// TIA Portal project "Automatizare_RT" (V17)

(* hardware
DEVICE "S7-300/ET200M station_1"  S7-300 station
   slot 0: "Rail_0"  Rail  6ES7 390-1***0-0AA0
   slot 1: "PS 307 5A_1"  PS 307 5A  6ES7 307-1EA00-0AA0
   slot 2: "PLC_1"  CPU 319-3 PN/DP  6ES7 318-3EL00-0AB0  V2.6
      slot 1: "MPI/DP interface_1"  X1
      slot 2: "DP interface_1"  X2
      slot 3: "PROFINET interface_1"  PN-IO
         slot 1: "Port_1"  Port
   slot 4: "DI 8/DO 8x24VDC/0.5A_1"  DI8/DO8 x 24VDC / 0.5A  6ES7 323-1BH01-0AA0
   slot 5: "DI 8/DO 8x24VDC/0.5A_2"  DI8/DO8 x 24VDC / 0.5A  6ES7 323-1BH01-0AA0
   slot 6: "AI 8x12BIT_1"  AI8 x 12 bits  6ES7 331-7KF02-0AB0
DEVICE "HMI_1"  KTP600 Basic color PN
   slot 0: "HMI_1"  KTP600 Basic color PN  6AV6 647-0AD11-3AX0  12.0.0.0
   slot 1: "HMI_RT_2"  KTP600 Basic color PN  6AV6 647-0AD11-3AX0  12.0.0.0
   slot 5: "HMI_1.IE_CP_1"  PROFINET Interface  12.0.0.0
      slot 1: "PROFINET Interface_1"  PROFINET Interface
         slot 1: "Port_1"  Port
DEVICE "PC-System_2"  SIMATIC PC station
   slot 0: "SIMATIC PC station"  Rail  SIMATIC PC-Station  V1.0
      slot 125: "Stationmanager"  Station_Manager  V6.0.4
   slot 1: "CP 1628_1"  CP 1628  6GK1 162-8AA00  V8.2.2
   slot 3: "HMI_RT_3"  WinCC RT Advanced  6AV2 104-0xxxx-xxxx  17.0.0.0
      slot 33792: "Computer interface"  Host interface
DEVICE "S7-1500/ET200MP station_1"  S7-1500 station
   slot 0: "Rail_0"  Rack  6ES7 590-1***0-0AA0
   slot 1: "PLC_2"  CPU 1518-4 PN/DP  6ES7 518-4AP00-0AB0  V2.9
      slot 3: "CPU display_1"  6ES7591-1BA00-0AA0
      slot 32768: "PROFINET interface_1"  X1
         slot 32769: "Port_1"  X1 P1
         slot 32770: "Port_2"  X1 P2
      slot 33024: "PROFINET interface_2"  X2
         slot 33025: "Port_1"  X2 P1
      slot 33280: "PROFINET interface GBIT_3"  X3
         slot 33281: "Port_1"  X3 P1
      slot 33536: "DP interface_1"  X4
      slot 34817: "Virtual CP interface port_1"  Virtual CP interface port  Virtual CP interface port
*)

// ===== PLC "PLC_1"  CPU 319-3 PN/DP =====

VAR_GLOBAL   // PLC tag table "Default tag table"
   "Pozitie_Incarcare" AT %Q1.6 : Bool;
   "Pozitie_Descarcare" AT %Q1.7 : Bool;
   "Status_Banda_1" AT %Q3.4 : Bool;
   "Mod_Operare" AT %Q3.5 : Bool;
   "Start/Stop" AT %Q3.6 : Bool;
   "Delimitare_Interval" AT %M100.0 : Bool;
   "10HzFcnTag" AT %M300.0 : Bool;
   "10Hz" AT %M300.1 : Bool;
   "ON/OFF" AT %M2.1 : Bool;
   "LOAD" AT %M2.4 : Bool;
   "Place_Box" AT %M2.6 : Bool;
   "TrigPozCutieCapatBanda1" AT %M200.1 : Bool;
   "5_Hz" AT %M500.1 : Bool;
   "10_Hz" AT %M500.0 : Bool;
   "1.25_Hz" AT %M500.4 : Bool;
   "0.5Hz" AT %M500.7 : Bool;
   "TrigPlaceBoxModAuto" AT %M3000.2 : Bool;
   "TrigVizCutieScurtaModAuto" AT %M3000.3 : Bool;
   "TrigAckLoadModAuto" AT %M3000.4 : Bool;
   "TrigPozCutie99AnimatieB1" AT %M3000.6 : Bool;
   "TrigPistonIncarcareA" AT %M400.0 : Bool;
   "TrigPistonIncarcareB" AT %M400.2 : Bool;
   "TrigPistonIncarcareC" AT %M400.4 : Bool;
   "QCounterRacire" AT %M600.0 : Bool;
   "QCounterIncalzire" AT %M600.1 : Bool;
   "2.5_Hz" AT %M500.2 : Bool;
   "TrigVizCutiePoz99CutieLung1" AT %M600.4 : Bool;
   "TrigGreutate100FCNCantar" AT %M800.0 : Bool;
   "TrigGreutate100FCNCantar2" AT %M800.1 : Bool;
   "TrigGreutate150FCNCantar" AT %M800.2 : Bool;
   "TrigGreutate150FCNCantar2" AT %M800.3 : Bool;
   "TrigPozCutie99CutieLung2" AT %M900.0 : Bool;
   "Tag_1" AT %M765.0 : Bool;
   "Tag_2" AT %M217.1 : Bool;
   "Tag_3" AT %M218.0 : Bool;
   "Tag_4" AT %M218.1 : Bool;
   "Tag_5" AT %M218.2 : Bool;
   "Tag_6" AT %M219.0 : Bool;
END_VAR

VAR_GLOBAL   // PLC tag table "Tab_tag_Motoare"
   "Motor_1_banda_1_DIST_Start_KL_FB" AT %Q0.0 : Bool;
   "Motor_1_banda_1_DIST_Start_K1_FB" AT %Q0.1 : Bool;
   "Motor_1_banda_1 _DIST_Start_K2_FB" AT %Q0.2 : Bool;
   "Motor_1_banda_1_LOC_Start_KL_FB" AT %Q0.3 : Bool;
   "Motro_1_banda_1_LOC_Start_K1_FB" AT %Q0.4 : Bool;
   "Motor_1_banda_1_LOC_Start_K2_FB" AT %Q0.5 : Bool;
   "Motor_2_banda_1_DIST_Start_KL_FB" AT %Q0.6 : Bool;
   "Motor_2_banda_1_DIST_Start_K1_FB" AT %Q0.7 : Bool;
   "Motor_2_banda_1 _DIST_Start_K2_FB" AT %Q1.0 : Bool;
   "Motor_2_banda_1_LOC_Start_KL_FB" AT %Q1.1 : Bool;
   "Motro_2_banda_1_LOC_Start_K1_FB" AT %Q1.2 : Bool;
   "Motor_2_banda_1_LOC_Start_K2_FB" AT %Q1.3 : Bool;
   "Motor_1_banda_1_Protectii_FB" AT %Q1.4 : Bool;
   "Motor_2_banda_1_Protectii_FB" AT %Q1.5 : Bool;
   "Motor_1_banda_1_DIST_Start_ON_KL" AT %Q2.0 : Bool;
   "Motor_1_banda_1_DIST_Start_ON_K1" AT %Q2.1 : Bool;
   "Motor_1_banda_1 _DIST_Start_ON_K2" AT %Q2.2 : Bool;
   "Motor_1_banda_1_LOC_Start_ON_KL" AT %Q2.3 : Bool;
   "Motro_1_banda_1_LOC_Start_ON_K1" AT %Q2.4 : Bool;
   "Motor_1_banda_1_LOC_Start_ON_K2" AT %Q2.5 : Bool;
   "Motor_2_banda_1_DIST_Start_ON_KL" AT %Q2.6 : Bool;
   "Motor_2_banda_1_DIST_Start_ON_K1" AT %Q2.7 : Bool;
   "Motor_2_banda_1 _DIST_Start_ON_K2" AT %Q3.0 : Bool;
   "Motor_2_banda_1_LOC_Start_ON_KL" AT %Q3.1 : Bool;
   "Motro_2_banda_1_LOC_Start_ON_K1" AT %Q3.2 : Bool;
   "Motor_2_banda_1_LOC_Start_ON_K2" AT %Q3.3 : Bool;
END_VAR

VAR_GLOBAL   // PLC tag table "Butoane"
   "Start" AT %I0.0 : Bool;
   "Stop" AT %I0.1 : Bool;
   "Emg_Stop" AT %I0.2 : Bool;
   "Man/Auto" AT %I0.3 : Bool;   // 0=manual/1=automat
END_VAR

VAR_GLOBAL   // PLC tag table "Tag_Animatii"
   "Poz_Cutie" AT %MW0 : Int;
   "Poz_Piston_1" AT %MW9 : Int;
   "Viz_Cutie_Cursa_Scurta" AT %M2.2 : Bool;
   "Viz_Cutie_Cursa_Lunga" AT %M2.3 : Bool;
   "Final_Cursa_Piston_1" AT %M2.5 : Bool;
   "Ecran_Stare_Descarcare" AT %M2.7 : Bool;   // Cand acesta devine 1 se face tranzitia la Statie Descarcare
END_VAR

// folder: Global Data/ DB

DATA_BLOCK "DB_general"   // DB2
{ S7_Optimized_Access := 'FALSE' }
VERSION : 0.1
   VAR
      Stare_Poz_Incarcare : Bool;
      Stare_Poz_Descarcare : Bool;
      Senzor_1_Incarcare : Bool;
      Senzor_2_Incarcare : Bool;
      Senzor_1_Descarcare : Bool;
      Senzor_2_Descarcare : Bool;
      Status_Banda_1 : Bool;
      Piston1_ON : Bool;
      Senzor_Prezenta_P1 : Bool;
      Btn_AKN_LOAD : Bool;
      Piston_1_In_Cursa : Bool;
      Poz_Piston_1 : Int;
      Poz_Cutie : Int;
      "Limita_Counter(50)" : Bool;
      Final_Cursa_Bile : Bool;
      Poz_Cutie_Bile : Int := 1;
      Status_Banda_2 : Bool;
      Inceput_Cursa_Bile : Int;
      Valoare : Int;
      Piston_1_Cursa_Completa : Int := 1;
      Piston_2_Cursa_Completa : Int := 1;
      zero_or_less : Bool;
      Poz_Max : Int := 25;
      Poz_Initiala : Int := 0;
      Max_Cursa_P1 : Bool;
      Max_Cursa_P2 : Bool;
      Max_Cursa_Banda : Bool;
      Piston_Incarcare : Int := 3;
      Piston_Incarcare_A : Int;
      Piston_Incarcare_B : Int;
      Piston_Incarcare_C : Int;
      Piston_Scrap : Int;
      Max_P_Incarcare : Bool;
      Auz_Volum_Ulei : Int;
      CondOptimePistoane : Bool;
      GreutateManual : Real;
      GreutateAutomata : Real;
      Procent_Toleranta : Real;
      TolerantaManual : Real;
      TolerantaAutomat : Real;
      Procent : Real;
      GreutateMinManual : Real;
      GreutateMaxManual : Real;
      GreutateMinAutomat : Real;
      GreutateMaxAutomat : Real;
      "100-P" : Real;
      "100+P" : Real;
   END_VAR
BEGIN
END_DATA_BLOCK

DATA_BLOCK "DB_RemoteAcces"   // DB6
{ S7_Optimized_Access := 'FALSE' }
VERSION : 0.1
   VAR
      EmgStopBtn : Bool;
      Stop : Bool;
      Start : Bool;
      "Manual/Auto" : Bool;
      "On/Off" : Bool;
      Remote : Bool;
      ControlEnable_Stop : Bool;
      ControlEnable_Start : Bool;
      "ControlEnable_Man/Auto" : Bool;
   END_VAR
BEGIN
END_DATA_BLOCK

DATA_BLOCK "Data_Control_En"   // DB14
{ S7_Optimized_Access := 'FALSE' }
VERSION : 0.1
   VAR
      Load_Enable : Bool;
      Destination_Enable : Bool;
      Manual_Enable : Bool;
   END_VAR
BEGIN
END_DATA_BLOCK

DATA_BLOCK "Template"   // DB16
{ S7_Optimized_Access := 'FALSE' }
VERSION : 0.1
   VAR
      Satie_Distribuire : Bool;
      Statie_Incarcare : Bool;
      Packets_Log : Bool;
      Hidraulic_Station : Bool;
      Errors : Bool;
      Home : Bool;
   END_VAR
BEGIN
END_DATA_BLOCK

DATA_BLOCK "DB_HMI"   // DB19
{ S7_Optimized_Access := 'FALSE' }
VERSION : 0.1
   VAR
      Locuri_A : Int := 3;
      Locuri_B : Int := 3;
      Locuri_C : Int := 3;
      A_Pressed : Bool;
      B_Pressed : Bool;
      C_Pressed : Bool;
      Cutie_Automata : Bool;
      Cutie_Manuala : Bool;
      Viz_Cutie_Scurta : Bool;
      Viz_Cutie_Lunga : Bool;
      Tip_Cutie_Lung : Int := 1;
      Tip_Cutie_Scurt : Int;
      LOAD : Int;
      Transport : Bool;
      "bool" : Bool;
      Viz_Cutie_Banda_1 : Bool;
      Ack_Load : Bool;
      Piston_1_Status : Int;
      Piston_2_Status : Int;
      Load_RDY : Bool;
      Viz_Cutie_A : Bool;
      Viz_Cutie_B : Bool;
      Viz_Cutie_C : Bool;
      Status_Piston_A : Int;
      Status_Piston_B : Int;
      Status_Piston_C : Int;
      LOAD_A : Bool;
      LOAD_B : Bool;
      LOAD_C : Bool;
      Status_Banda_Bile : Int;
      Sageata_Deplasare_Banda_Bile : Bool;
      Temp_Ulei : Int := 0;
      Temp_Ulei_Min : Int;
      Temp_Ulei_Max : Int;
      Volum_Ulei : Int := 40;
      Add_Ulei : Bool;
      Sub_Ulei : Bool;
      Start_System : Bool;
      Racire_Ulei : Bool;
      Incalzire_Ulei : Bool;
      Oricare_Piston : Bool;
      Set_T0 : Bool;
      Set_T50 : Bool;
      START_SIM : Bool;
      BTN_LOAD : Bool;
      "Status_Incalzire/Racire_Ulei" : Int;
      "Viz_Cutie_Man/Auto" : Int;
      Ventilator_Rece : Int;
      Ventilator_Cald : Int;
      Viz_Platforma_Libera : Bool;
      Greutate : Real;
      Nr_runuri : Int;
      rest_runuri : Int;
      Nr_Run : DInt;
      Rest_Run : DInt;
      Shift_Details : Int;
      Packets_Param : Int;
      MaxLoad_A : Int;
      MaxLoad_B : Int;
      MaxLoad_C : Int;
      Cantitate_A : Int;
      Cantitate_B : Int;
      Cantitat_C : Int;
      Total_Packets : Int;
      Pachete_Schimb1 : Int;
      Pachete_Schimb2 : Int;
      Pachete_Schimb3 : Int;
      Cooling_Param : Bool;
      Temp_Max : Int := 40;
      Temp_Min : Int := 30;
      Temp_Optim : Int := 35;
      Total_Weight_A : Real;
      Total_Weight_B : Real;
      Total_Weight_C : Real;
      Cantitate_Loaded_A : Int;
      Cantitate_Loaded_B : Int;
      Cantitate_Loaded_C : Int;
      Detalii_Truck_A : Bool;
      Detalii_Truck_B : Bool;
      Detalii_Truck_C : Bool;
      Status_Piston_3 : Int;
      Eng : Bool;
      Weight_A : Real;
      Weight_B : Real;
      Weight_C : Real;
      Ger : Bool;
   END_VAR
BEGIN
END_DATA_BLOCK

DATA_BLOCK "DB_Butoane"   // DB33
{ S7_Optimized_Access := 'FALSE' }
VERSION : 0.1
   VAR
      Emg_Stop : Bool;
      Start : Bool;
      Stop : Bool;
      "Man/Auto" : Bool;
   END_VAR
BEGIN
END_DATA_BLOCK

DATA_BLOCK "DB_Tip_Cutie"   // DB37
{ S7_Optimized_Access := 'FALSE' }
VERSION : 0.1
   VAR
      GreutateCutie : Real;
      IntersectieInterval : Int;
      TipCutie : Bool;
      VizTipCutie : Bool;
      RebutLbl : Bool;
      BoxStatus : Bool;
      Scrap : Int;
   END_VAR
BEGIN
END_DATA_BLOCK

DATA_BLOCK "DB_SIM"   // DB40
{ S7_Optimized_Access := 'FALSE' }
VERSION : 0.1
   VAR
      Place_Box : Bool;
      Ack_Load : Bool;
      Load : Bool;
      Ack_Load_Pressed : Bool;
      BTN_RESET : Bool;
      Btn_Start_Sim : Bool;
   END_VAR
BEGIN
END_DATA_BLOCK

DATA_BLOCK "DB_ControlEnable"   // DB45
{ S7_Optimized_Access := 'FALSE' }
VERSION : 0.1
   VAR
      ControlEnable_Btn_A : Bool;
      ControlEnable_Btn_B : Bool;
      ControlEnable_Btn_C : Bool;
      ControlEnable_Btn_Load : Bool;
      ControlEnable_Btn_ACKLoad : Bool;
      ControlEnable_StartSim : Bool;
      ControlEnable_Btn_PlaceBox : Bool;
      StatusLoadBtn : Int;
      StatusACKBtn : Int;
      StatusPlaceBoxBtn : Int;
   END_VAR
BEGIN
END_DATA_BLOCK

DATA_BLOCK "DB_Alarme"   // DB46
{ S7_Optimized_Access := 'FALSE' }
VERSION : 0.1
   VAR
      Emg_Stop : Int;
   END_VAR
BEGIN
END_DATA_BLOCK

DATA_BLOCK "DB_Tranzitii"   // DB47
{ S7_Optimized_Access := 'FALSE' }
VERSION : 0.1
   VAR
      VizCutieStart : Bool;
      "Tip_Cutie_Man/Auto_Start" : Int;
      VizCutieEnd : Bool;
      "TipCutieMan/Auto_End" : Int;
      Viz_CutieScrapP3 : Bool;
      test : Bool;
   END_VAR
BEGIN
END_DATA_BLOCK

DATA_BLOCK "Errors"   // DB51
{ S7_Optimized_Access := 'FALSE' }
VERSION : 0.1
   VAR
      "Error information OB121" : Struct
         "Fault indentifier" : Byte;
      END_STRUCT;
   END_VAR
BEGIN
END_DATA_BLOCK

// folder: Global Data/Functii

DATA_BLOCK "10HzFcnDB"   // DB3
{ S7_Optimized_Access := 'FALSE' }
VERSION : 0.1
// stored: InstanceOfName 10HzFcn
"10HzFcn"
BEGIN
END_DATA_BLOCK

DATA_BLOCK "DB_InsertCutieTrigger"   // DB5
{ S7_Optimized_Access := 'FALSE' }
VERSION : 0.1
// stored: InstanceOfName InsertCutieTrigger
"InsertCutieTrigger"
BEGIN
END_DATA_BLOCK

DATA_BLOCK "Tip_Cutie_DB"   // DB21
{ S7_Optimized_Access := 'FALSE' }
VERSION : 0.1
// stored: InstanceOfName Tip_Cutie
"Tip_Cutie"
BEGIN
END_DATA_BLOCK

DATA_BLOCK "DB_ModAuto"   // DB42
{ S7_Optimized_Access := 'FALSE' }
VERSION : 0.1
// stored: InstanceOfName ModAuto
"ModAuto"
BEGIN
END_DATA_BLOCK

// folder: Hidraulic/DB

DATA_BLOCK "DB_Status_Motoare"   // DB25
{ S7_Optimized_Access := 'FALSE' }
VERSION : 0.1
   VAR
      Motor_1 : Int;
      Motor_2 : Int;
      Motor_3 : Int;
   END_VAR
BEGIN
END_DATA_BLOCK

DATA_BLOCK "DB_Status_Pistoane"   // DB26
{ S7_Optimized_Access := 'FALSE' }
VERSION : 0.1
   VAR
      Status_Piston_1 : Int;
      Status_Pison_2 : Int;
      Status_Piston_A : Int;
      Status_Piston_B : Int;
      Status_Piston_C : Int;
   END_VAR
BEGIN
END_DATA_BLOCK

DATA_BLOCK "DB_Inspect_Pistoane"   // DB34
{ S7_Optimized_Access := 'FALSE' }
VERSION : 0.1
   VAR
      Piston_1 : Bool;
      Piston_2 : Bool;
      Piston_A : Bool;
      Piston_B : Bool;
      Piston_C : Bool;
      Inspect_Pistoane : Bool;
      Presiune_1 : Int := 3;
      Presiune_2 : Int := 3;
      Presiune_A : Int := 3;
      Presiune_B : Int := 3;
      Presiune_C : Int := 3;
      Presiune_Upper_2 : Int := 5;
      Presiune_Upper_1 : Int := 4;
      Presiune_Lower_1 : Int := 2;
      Presiune_Lower_2 : Int := 1;
      PompaPrincipala : Int := 2;
      Pompa1 : Int := 2;
      Pompa2 : Int := 2;
      PompaA : Int := 2;
      PompaB : Int := 2;
      PompaC : Int := 2;
      TrigPiston1 : Bool;
      TrigPiston2 : Bool;
      TrigPistonA : Bool;
      TrigPistonB : Bool;
      TrigPistonC : Bool;
      CutP1 : Bool;
      StatusPump1 : Int := 1;
      StatusPump2 : Int := 1;
      StatusPumpA : Int := 1;
      StatusPumpB : Int := 1;
      StatusPumpC : Int := 1;
   END_VAR
BEGIN
END_DATA_BLOCK

// folder: Statie Distribuire/Animatii

DATA_BLOCK "Animatie_Banda_1_DB"   // DB13
{ S7_Optimized_Access := 'FALSE' }
VERSION : 0.1
// stored: InstanceOfName Animatie_Banda_1
"Animatie_Banda_1"
BEGIN
END_DATA_BLOCK

DATA_BLOCK "Animatie_Piston_1_DB"   // DB18
{ S7_Optimized_Access := 'FALSE' }
VERSION : 0.1
// stored: InstanceOfName Animatie_Piston_1
"Animatie_Piston_1"
BEGIN
END_DATA_BLOCK

DATA_BLOCK "Piston_Cursa_Completa_DB"   // DB27
{ S7_Optimized_Access := 'FALSE' }
VERSION : 0.1
// stored: InstanceOfName Piston_1_Cursa_Completa
"Piston_1_Cursa_Completa"
BEGIN
END_DATA_BLOCK

DATA_BLOCK "Piston_2_Cursa_Completa_DB"   // DB28
{ S7_Optimized_Access := 'FALSE' }
VERSION : 0.1
// stored: InstanceOfName Piston_2_Cursa_Completa
"Piston_2_Cursa_Completa"
BEGIN
END_DATA_BLOCK

DATA_BLOCK "DB_TranzitieBanda1-Graph"   // DB50
{ S7_Optimized_Access := 'FALSE' }
VERSION : 0.1
// stored: InstanceOfName TranzitieBanda1-Graph
"TranzitieBanda1-Graph"
BEGIN
END_DATA_BLOCK

// folder: Statie Distribuire/Functii

DATA_BLOCK "DB_Verificare_Poz_StartSec"   // DB4
{ S7_Optimized_Access := 'FALSE' }
VERSION : 0.1
// stored: InstanceOfName Verificare_Poz_StartSec
"Verificare_Poz_StartSec"
BEGIN
END_DATA_BLOCK

DATA_BLOCK "Cantar_DB"   // DB7
{ S7_Optimized_Access := 'FALSE' }
VERSION : 0.1
// stored: InstanceOfName Cantar
"Cantar"
BEGIN
END_DATA_BLOCK

DATA_BLOCK "Banda_1_DB"   // DB8
{ S7_Optimized_Access := 'FALSE' }
VERSION : 0.1
// stored: InstanceOfName Banda_1
"Banda_1"
BEGIN
END_DATA_BLOCK

DATA_BLOCK "Verificare_Poz_Capat_DB"   // DB12
{ S7_Optimized_Access := 'FALSE' }
VERSION : 0.1
// stored: InstanceOfName Verificare_Poz_StartSec
"Verificare_Poz_StartSec"
BEGIN
END_DATA_BLOCK

// folder: Statie Incarcare/Animatii

DATA_BLOCK "DB_Vizibilitati_Platforme/Colete"   // DB1
{ S7_Optimized_Access := 'FALSE' }
VERSION : 0.1
   VAR
      Platforma_A : Bool;
      Platforma_B : Bool;
      Platforma_C : Bool;
      Colet_A : Bool;
      Colet_B : Bool;
      Colet_C : Bool;
      Rebut : Bool;
      Colet_Rebut : Bool;
      Platforma_Rebut : Bool;
   END_VAR
BEGIN
END_DATA_BLOCK

DATA_BLOCK "Animatie_Banda_Bile_DB"   // DB24
{ S7_Optimized_Access := 'FALSE' }
VERSION : 0.1
// stored: InstanceOfName Animatie_Banda_Bile
"Animatie_Banda_Bile"
BEGIN
END_DATA_BLOCK

DATA_BLOCK "Piston_Incarcare_DB"   // DB32
{ S7_Optimized_Access := 'FALSE' }
VERSION : 0.1
// stored: InstanceOfName Piston_Incarcare
"Piston_Incarcare"
BEGIN
END_DATA_BLOCK

// folder: Statie Incarcare/Functii

DATA_BLOCK "Banda_Bile_DB"   // DB23
{ S7_Optimized_Access := 'FALSE' }
VERSION : 0.1
// stored: InstanceOfName Banda_Bile
"Banda_Bile"
BEGIN
END_DATA_BLOCK

DATA_BLOCK "DB_Banda_Bile_Poz_Reset"   // DB41
{ S7_Optimized_Access := 'FALSE' }
VERSION : 0.1
   VAR
      "Counter" : Int;
   END_VAR
BEGIN
END_DATA_BLOCK

// folder: Statie Retur

DATA_BLOCK "DB_Banda3"   // DB49
{ S7_Optimized_Access := 'FALSE' }
VERSION : 0.1
   VAR
      Poz_Banda3 : Int;
      Viz_CutieBanda3 : Bool;
      AckScrap : Bool;
   END_VAR
BEGIN
END_DATA_BLOCK

// folder: (top level)

ORGANIZATION_BLOCK "Main"   // OB1, FBD
TITLE = "Main Program Sweep (Cycle)"
{ S7_Optimized_Access := 'FALSE' }
VERSION : 0.1
   VAR_TEMP
      OB1_EV_CLASS : Byte;   // Bits 0-3 = 1 (Coming event), Bits 4-7 = 1 (Event class 1)
      OB1_SCAN_1 : Byte;   // 1 (Cold restart scan 1 of OB 1), 3 (Scan 2-n of OB 1)
      OB1_PRIORITY : Byte;   // Priority of OB Execution
      OB1_OB_NUMBR : Byte;   // 1 (Organization block 1, OB1)
      OB1_RESERVED_1 : Byte;   // Reserved for system
      OB1_RESERVED_2 : Byte;   // Reserved for system
      OB1_PREV_CYCLE : Int;   // Cycle time of previous OB1 scan (milliseconds)
      OB1_MIN_CYCLE : Int;   // Minimum cycle time of OB1 (milliseconds)
      OB1_MAX_CYCLE : Int;   // Maximum cycle time of OB1 (milliseconds)
      OB1_DATE_TIME : Date_And_Time;   // Date and time OB1 started
   END_VAR
BEGIN

REGION Network 1: Verif pozitie capat incarcare / Check_Pos_Loadhead
   // Verifi stare pozitie incarcare / Überprüfen Sie den Status der Ladeposition
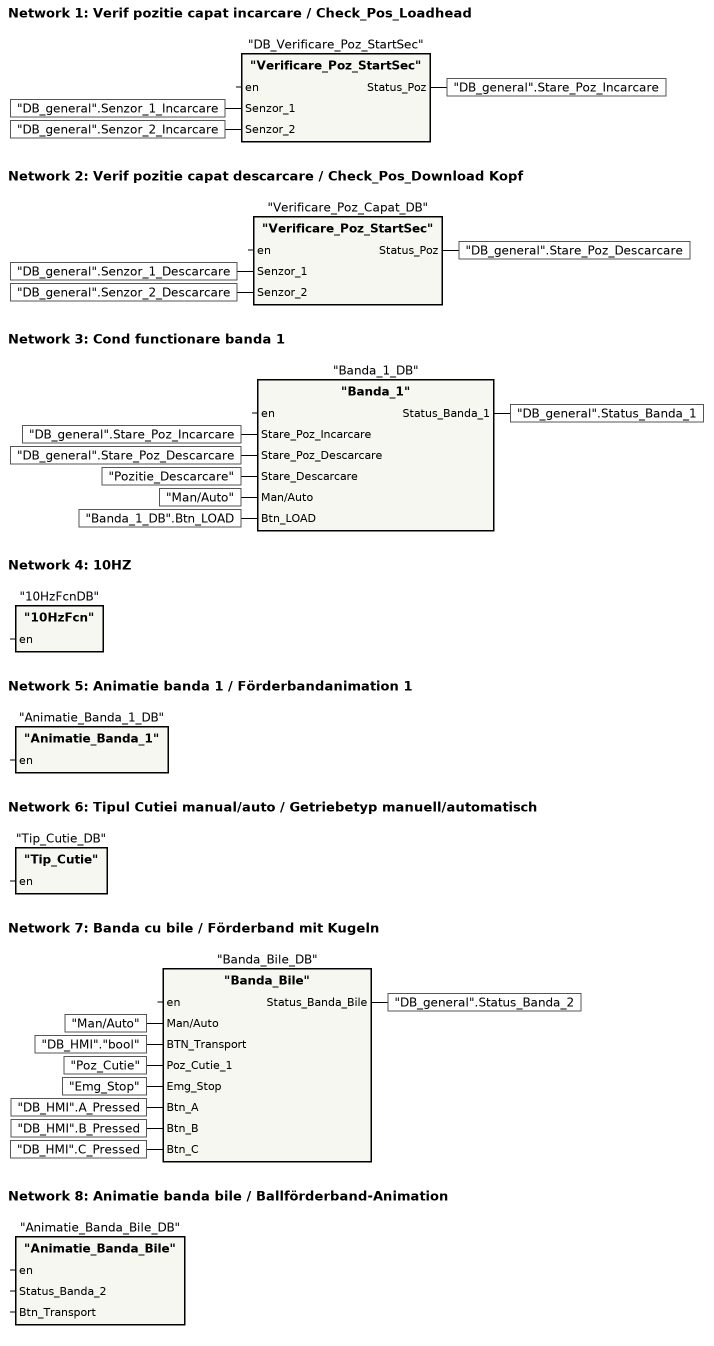
   "DB_Verificare_Poz_StartSec"(Senzor_1 := "DB_general".Senzor_1_Incarcare,   // "Verificare_Poz_StartSec"
                           Senzor_2 := "DB_general".Senzor_2_Incarcare,
                           Status_Poz => "DB_general".Stare_Poz_Incarcare);
END_REGION

REGION Network 2: Verif pozitie capat descarcare / Check_Pos_Download Kopf
   // Überprüfen Sie den Status der Ladeposition / Überprüfen Sie den Status der Anzahlung
   "Verificare_Poz_Capat_DB"(Senzor_1 := "DB_general".Senzor_1_Descarcare,   // "Verificare_Poz_StartSec"
                           Senzor_2 := "DB_general".Senzor_2_Descarcare,
                           Status_Poz => "DB_general".Stare_Poz_Descarcare);
END_REGION

REGION Network 3: Cond functionare banda 1
   // Banda 1 / Förderband 1
   "Banda_1_DB"(Stare_Poz_Incarcare := "DB_general".Stare_Poz_Incarcare,   // "Banda_1"
                Stare_Poz_Descarcare := "DB_general".Stare_Poz_Descarcare,
                Stare_Descarcare := "Pozitie_Descarcare",
                "Man/Auto" := "Man/Auto",
                Btn_LOAD := "Banda_1_DB".Btn_LOAD,
                Status_Banda_1 => "DB_general".Status_Banda_1);
END_REGION

REGION Network 4: 10HZ
   "10HzFcnDB"();   // "10HzFcn"
END_REGION

REGION Network 5: Animatie banda 1 / Förderbandanimation 1
   "Animatie_Banda_1_DB"();   // "Animatie_Banda_1"
END_REGION

REGION Network 6: Tipul Cutiei manual/auto / Getriebetyp manuell/automatisch
   "Tip_Cutie_DB"();   // "Tip_Cutie"
END_REGION

REGION Network 7: Banda cu bile / Förderband mit Kugeln
   "Banda_Bile_DB"("Man/Auto" := "Man/Auto",   // "Banda_Bile"
                   BTN_Transport := "DB_HMI"."bool",
                   Poz_Cutie_1 := "Poz_Cutie",
                   Emg_Stop := "Emg_Stop",
                   Btn_A := "DB_HMI".A_Pressed,
                   Btn_B := "DB_HMI".B_Pressed,
                   Btn_C := "DB_HMI".C_Pressed,
                   Status_Banda_Bile => "DB_general".Status_Banda_2);
END_REGION

REGION Network 8: Animatie banda bile / Ballförderband-Animation
   "Animatie_Banda_Bile_DB"();   // "Animatie_Banda_Bile"
END_REGION

REGION Network 9: Cursa completa a pistonului 1 / Voller Hub von Kolben 1
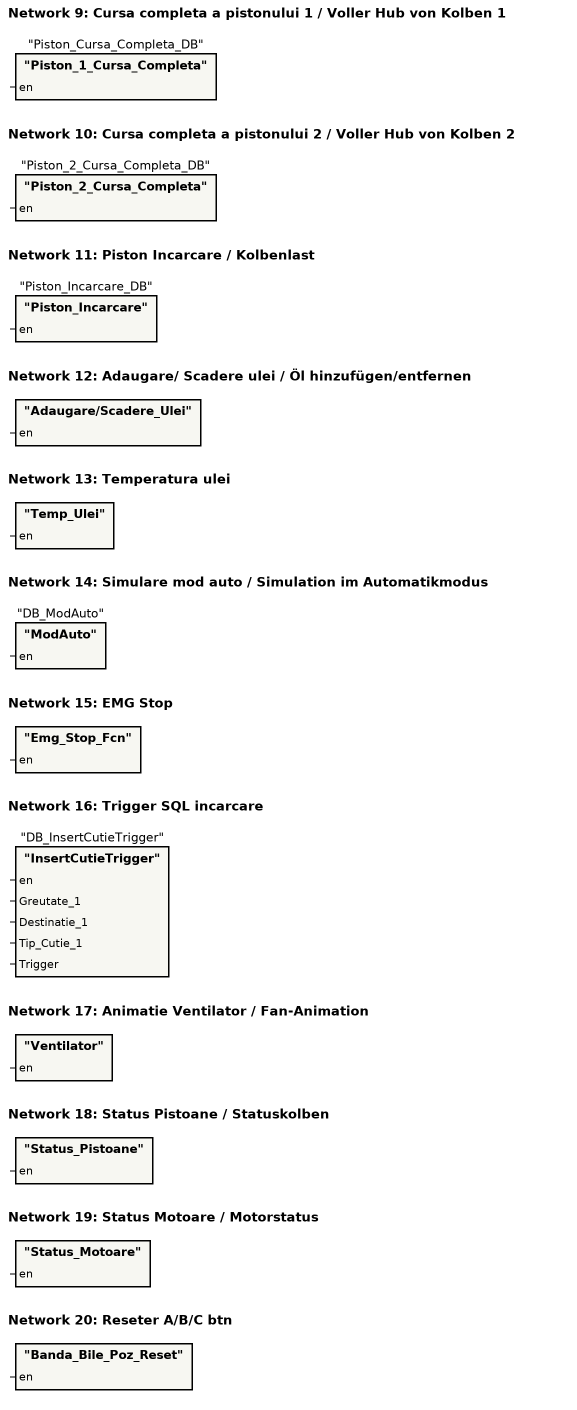
   "Piston_Cursa_Completa_DB"();   // "Piston_1_Cursa_Completa"
END_REGION

REGION Network 10: Cursa completa a pistonului 2 / Voller Hub von Kolben 2
   "Piston_2_Cursa_Completa_DB"();   // "Piston_2_Cursa_Completa"
END_REGION

REGION Network 11: Piston Incarcare / Kolbenlast
   "Piston_Incarcare_DB"();   // "Piston_Incarcare"
END_REGION

REGION Network 12: Adaugare/ Scadere ulei / Öl hinzufügen/entfernen
   "Adaugare/Scadere_Ulei"();
END_REGION

REGION Network 13: Temperatura ulei
   "Temp_Ulei"();
END_REGION

REGION Network 14: Simulare mod auto / Simulation im Automatikmodus
   "DB_ModAuto"();   // "ModAuto"
END_REGION

REGION Network 15: EMG Stop
   "Emg_Stop_Fcn"();
END_REGION

REGION Network 16: Trigger SQL incarcare
   "DB_InsertCutieTrigger"();   // "InsertCutieTrigger"
END_REGION

REGION Network 17: Animatie Ventilator / Fan-Animation
   "Ventilator"();
END_REGION

REGION Network 18: Status Pistoane / Statuskolben
   // 0-EROARE
   // 1-FUNCTIONARE
   // 2-STOP
   "Status_Pistoane"();
END_REGION

REGION Network 19: Status Motoare / Motorstatus
   // 0-EROARE
   // 1-FUNCTIONARE
   // 2-STOP
   "Status_Motoare"();
END_REGION

REGION Network 20: Reseter A/B/C btn
   "Banda_Bile_Poz_Reset"();
END_REGION

REGION Network 21: Tranzitii cutie pe banda transport 1-Graph / Kastenübergänge am Förderband 1
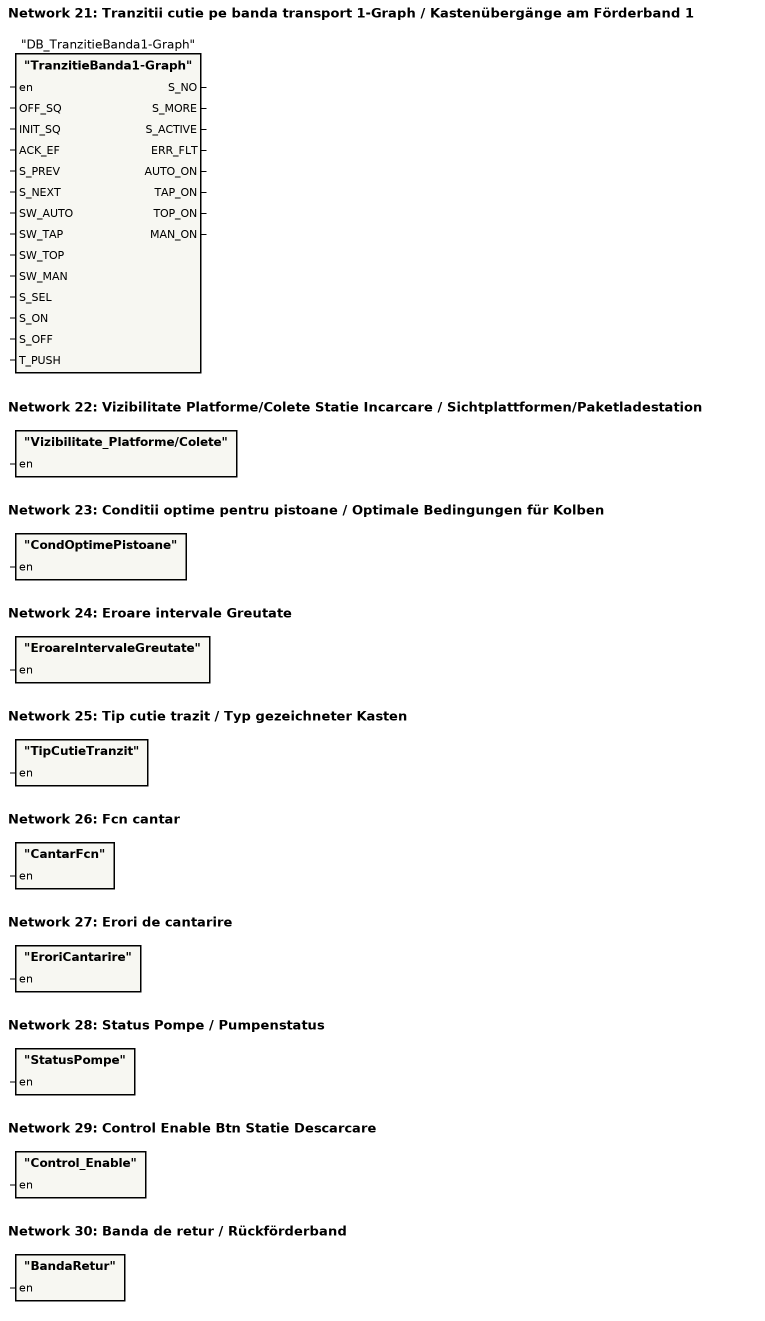
   "DB_TranzitieBanda1-Graph"();   // "TranzitieBanda1-Graph"
END_REGION

REGION Network 22: Vizibilitate Platforme/Colete Statie Incarcare / Sichtplattformen/Paketladestation
   "Vizibilitate_Platforme/Colete"();
END_REGION

REGION Network 23: Conditii optime pentru pistoane / Optimale Bedingungen für Kolben
   "CondOptimePistoane"();
END_REGION

REGION Network 24: Eroare intervale Greutate
   "EroareIntervaleGreutate"();
END_REGION

REGION Network 25: Tip cutie trazit / Typ gezeichneter Kasten
   "TipCutieTranzit"();
END_REGION

REGION Network 26: Fcn cantar
   "CantarFcn"();
END_REGION

REGION Network 27: Erori de cantarire
   "EroriCantarire"();
END_REGION

REGION Network 28: Status Pompe / Pumpenstatus
   "StatusPompe"();
END_REGION

REGION Network 29: Control Enable Btn Statie Descarcare
   "Control_Enable"();
END_REGION

REGION Network 30: Banda de retur / Rückförderband
   "BandaRetur"();
END_REGION

REGION Network 31: Consola Comanda
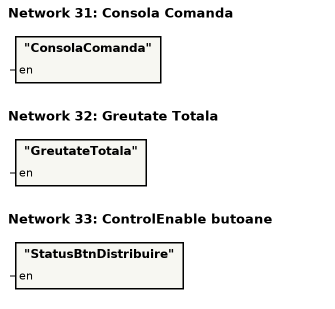
   "ConsolaComanda"();
END_REGION

REGION Network 32: Greutate Totala
   "GreutateTotala"();
END_REGION

REGION Network 33: ControlEnable butoane
   "StatusBtnDistribuire"();
END_REGION
END_ORGANIZATION_BLOCK

ORGANIZATION_BLOCK "PROG_ERR"   // OB121, FBD
TITLE = "Programming Error"
{ S7_Optimized_Access := 'FALSE' }
VERSION : 0.1
   VAR_TEMP
      OB121_EV_CLASS : Byte;   // 16#25, Event class 2, Entering event state, Internal fault event
      OB121_SW_FLT : Byte;   // 16#XX Software programming fault
      OB121_PRIORITY : Byte;   // Priority of OB Execution
      OB121_OB_NUMBR : Byte;   // 121 (Organization block 121, OB121)
      OB121_BLK_TYPE : Byte;   // 16#88/8A/8B/8C/8E Type of block fault occured in
      OB121_RESERVED_1 : Byte;   // Reserved for system
      OB121_FLT_REG : Word;   // 16#XX Specific register that caused fault
      OB121_BLK_NUM : Word;   // Number of block that programming fault occured in
      OB121_PRG_ADDR : Word;   // Address in block where programming fault occured
      OB121_DATE_TIME : Date_And_Time;   // Date and time OB121 started
   END_VAR
BEGIN
END_ORGANIZATION_BLOCK

// folder: Global Data/Functii

FUNCTION_BLOCK "10HzFcn"   // FB1, LAD
{ S7_Optimized_Access := 'FALSE' }
VERSION : 0.1
   VAR_TEMP
      increment : Bool;
   END_VAR
BEGIN

REGION Network 1
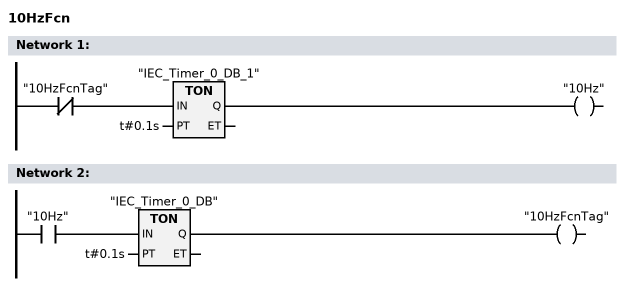
   "IEC_Timer_0_DB_1".TON(IN := NOT "10HzFcnTag", PT := t#0.1s);
   "10Hz" := "IEC_Timer_0_DB_1".Q;
END_REGION

REGION Network 2
   "IEC_Timer_0_DB".TON(IN := "10Hz", PT := t#0.1s);
   "10HzFcnTag" := "IEC_Timer_0_DB".Q;
END_REGION
END_FUNCTION_BLOCK

FUNCTION_BLOCK "InsertCutieTrigger"   // FB5, SCL
{ S7_Optimized_Access := 'FALSE' }
VERSION : 0.1
   VAR_INPUT
      Greutate_1 : Int;
      Destinatie_1 : Int;
      Tip_Cutie_1 : Int;
   END_VAR
   VAR_IN_OUT
      Trigger : Bool;
   END_VAR
   VAR
      Readytolog : Bool;
      Destinatie_Pachet : Int;
      Greutate_Pachet : Int;
      Tip_Cutie_Pachet : Int;
   END_VAR
BEGIN
   IF #Trigger = TRUE THEN


       #Greutate_Pachet := #Greutate_1;
       #Tip_Cutie_Pachet := #Tip_Cutie_1;
       #Destinatie_Pachet := #Destinatie_1;


       #Readytolog := TRUE;
       #Trigger := false;
   END_IF;
END_FUNCTION_BLOCK

FUNCTION_BLOCK "Tip_Cutie"   // FB14, LAD
{ S7_Optimized_Access := 'FALSE' }
VERSION : 0.1
BEGIN

REGION Network 1
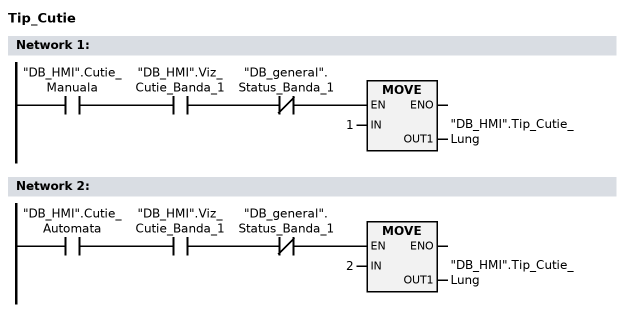
   RUNG wire#powerrail
      Contact( "DB_HMI".Cutie_Manuala )
      Contact( "DB_HMI".Viz_Cutie_Banda_1 )
      I_Contact( "DB_general".Status_Banda_1 )
      { S7_GenerateENO := "TRUE" } Move(in := 1, out1 => "DB_HMI".Tip_Cutie_Lung)
   END_RUNG
   // the same network as SCL:
   IF "DB_HMI".Cutie_Manuala AND "DB_HMI".Viz_Cutie_Banda_1 AND NOT "DB_general".Status_Banda_1 THEN
       "DB_HMI".Tip_Cutie_Lung := 1;
   END_IF;
END_REGION

REGION Network 2
   RUNG wire#powerrail
      Contact( "DB_HMI".Cutie_Automata )
      Contact( "DB_HMI".Viz_Cutie_Banda_1 )
      I_Contact( "DB_general".Status_Banda_1 )
      { S7_GenerateENO := "TRUE" } Move(in := 2, out1 => "DB_HMI".Tip_Cutie_Lung)
   END_RUNG
   // the same network as SCL:
   IF "DB_HMI".Cutie_Automata AND "DB_HMI".Viz_Cutie_Banda_1 AND NOT "DB_general".Status_Banda_1 THEN
       "DB_HMI".Tip_Cutie_Lung := 2;
   END_IF;
END_REGION
END_FUNCTION_BLOCK

FUNCTION_BLOCK "ModAuto"   // FB21, LAD
{ S7_Optimized_Access := 'FALSE' }
VERSION : 0.1
   VAR_TEMP   // added for the SCL form of the ladder/FBD networks
      _w1 : Bool;
      _w2 : Bool;
      _w3 : Bool;
      _w4 : Bool;
      _w5 : Bool;
      _w6 : Bool;
      _w7 : Bool;
      _w8 : Bool;
      _w9 : Bool;
   END_VAR
BEGIN

REGION Network 1
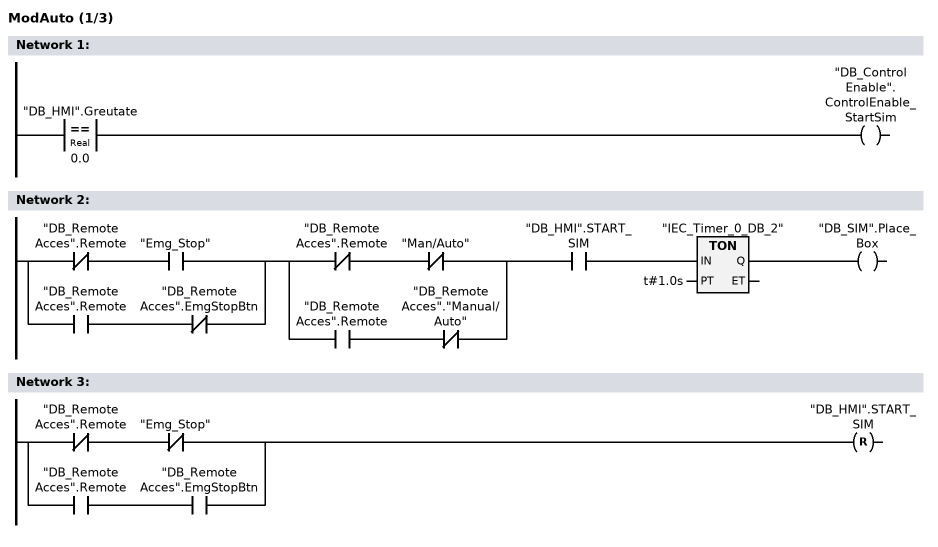
   RUNG wire#powerrail
      { S7_Templates := "SrcType := Real" } EQ_Contact(in1 := "DB_HMI".Greutate, in2 := 0.0)
      Coil( "DB_ControlEnable".ControlEnable_StartSim )
   END_RUNG
   // the same network as SCL:
   "DB_ControlEnable".ControlEnable_StartSim := "DB_HMI".Greutate = 0.0;
END_REGION

REGION Network 2
   "IEC_Timer_0_DB_2".TON(IN := ((NOT "DB_RemoteAcces".Remote AND "Emg_Stop") OR ("DB_RemoteAcces".Remote AND NOT "DB_RemoteAcces".EmgStopBtn)) AND ((NOT "DB_RemoteAcces".Remote AND NOT "Man/Auto") OR ("DB_RemoteAcces".Remote AND NOT "DB_RemoteAcces"."Manual/Auto")) AND "DB_HMI".START_SIM,
                          PT := t#1.0s);
   "DB_SIM".Place_Box := "IEC_Timer_0_DB_2".Q;
END_REGION

REGION Network 3
   RUNG wire#powerrail
      I_Contact( "DB_RemoteAcces".Remote )
      I_Contact( "Emg_Stop" )
      wire#w1
      R_Coil( "DB_HMI".START_SIM )
   END_RUNG
   RUNG wire#powerrail
      Contact( "DB_RemoteAcces".Remote )
      Contact( "DB_RemoteAcces".EmgStopBtn )
   END_RUNG wire#w1
   // the same network as SCL:
   IF (NOT "DB_RemoteAcces".Remote AND NOT "Emg_Stop") OR ("DB_RemoteAcces".Remote AND "DB_RemoteAcces".EmgStopBtn) THEN
       "DB_HMI".START_SIM := FALSE;
   END_IF;
END_REGION

REGION Network 4